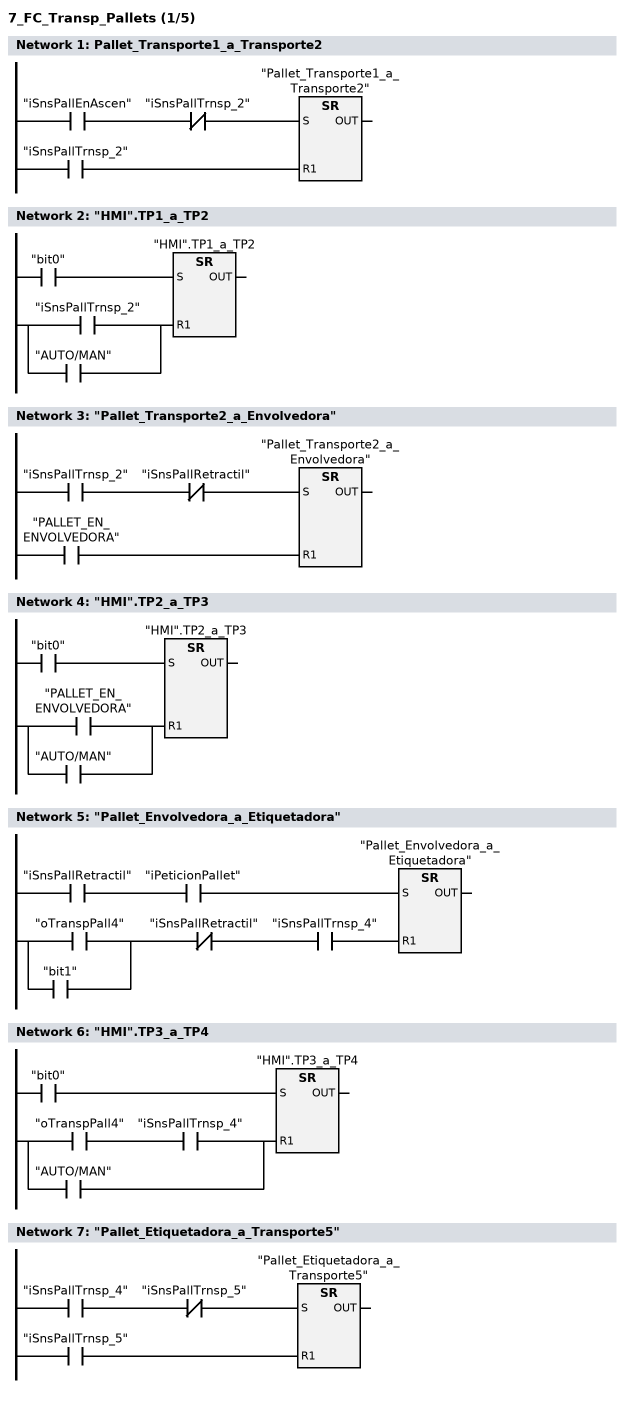
   RUNG wire#powerrail
      Contact( "iSnsPallEnAscen" )
      I_Contact( "iSnsPallTrnsp_2" )
      S_SR(operand := "Pallet_Transporte1_a_Transporte2", r1 := wire#w1)
   END_RUNG
   RUNG wire#powerrail
      Contact( "iSnsPallTrnsp_2" )
   END_RUNG wire#w1
   // the same network as SCL:
   IF "iSnsPallEnAscen" AND NOT "iSnsPallTrnsp_2" THEN
       "Pallet_Transporte1_a_Transporte2" := TRUE;   // SR flip-flop
   END_IF;
   IF "iSnsPallTrnsp_2" THEN "Pallet_Transporte1_a_Transporte2" := FALSE; END_IF;
END_REGION

REGION Network 2: "HMI".TP1_a_TP2
   RUNG wire#powerrail
      Contact( "bit0" )
      S_SR(operand := "HMI".TP1_a_TP2, r1 := wire#w1)
   END_RUNG
   RUNG wire#powerrail
      Contact( "iSnsPallTrnsp_2" )
   END_RUNG wire#w1
   RUNG wire#powerrail
      Contact( "AUTO/MAN" )
   END_RUNG wire#w1
   // the same network as SCL:
   IF "bit0" THEN
       "HMI".TP1_a_TP2 := TRUE;   // SR flip-flop
   END_IF;
   IF "iSnsPallTrnsp_2" OR "AUTO/MAN" THEN "HMI".TP1_a_TP2 := FALSE; END_IF;
END_REGION

REGION Network 3: "Pallet_Transporte2_a_Envolvedora"
   RUNG wire#powerrail
      Contact( "iSnsPallTrnsp_2" )
      I_Contact( "iSnsPallRetractil" )
      S_SR(operand := "Pallet_Transporte2_a_Envolvedora", r1 := wire#w1)
   END_RUNG
   RUNG wire#powerrail
      Contact( "PALLET_EN_ENVOLVEDORA" )
   END_RUNG wire#w1
   // the same network as SCL:
   IF "iSnsPallTrnsp_2" AND NOT "iSnsPallRetractil" THEN
       "Pallet_Transporte2_a_Envolvedora" := TRUE;   // SR flip-flop
   END_IF;
   IF "PALLET_EN_ENVOLVEDORA" THEN "Pallet_Transporte2_a_Envolvedora" := FALSE; END_IF;
END_REGION

REGION Network 4: "HMI".TP2_a_TP3
   RUNG wire#powerrail
      Contact( "bit0" )
      S_SR(operand := "HMI".TP2_a_TP3, r1 := wire#w1)
   END_RUNG
   RUNG wire#powerrail
      Contact( "PALLET_EN_ENVOLVEDORA" )
   END_RUNG wire#w1
   RUNG wire#powerrail
      Contact( "AUTO/MAN" )
   END_RUNG wire#w1
   // the same network as SCL:
   IF "bit0" THEN
       "HMI".TP2_a_TP3 := TRUE;   // SR flip-flop
   END_IF;
   IF "PALLET_EN_ENVOLVEDORA" OR "AUTO/MAN" THEN "HMI".TP2_a_TP3 := FALSE; END_IF;
END_REGION

REGION Network 5: "Pallet_Envolvedora_a_Etiquetadora"
   RUNG wire#powerrail
      Contact( "iSnsPallRetractil" )
      Contact( "iPeticionPallet" )
      S_SR(operand := "Pallet_Envolvedora_a_Etiquetadora", r1 := wire#w2)
   END_RUNG
   RUNG wire#powerrail
      Contact( "oTranspPall4" )
      wire#w1
      I_Contact( "iSnsPallRetractil" )
      Contact( "iSnsPallTrnsp_4" )
   END_RUNG wire#w2
   RUNG wire#powerrail
      Contact( "bit1" )
   END_RUNG wire#w1
   // the same network as SCL:
   IF "iSnsPallRetractil" AND "iPeticionPallet" THEN
       "Pallet_Envolvedora_a_Etiquetadora" := TRUE;   // SR flip-flop
   END_IF;
   IF ("oTranspPall4" OR "bit1") AND NOT "iSnsPallRetractil" AND "iSnsPallTrnsp_4" THEN
       "Pallet_Envolvedora_a_Etiquetadora" := FALSE;
   END_IF;
END_REGION

REGION Network 6: "HMI".TP3_a_TP4
   RUNG wire#powerrail
      Contact( "bit0" )
      S_SR(operand := "HMI".TP3_a_TP4, r1 := wire#w1)
   END_RUNG
   RUNG wire#powerrail
      Contact( "oTranspPall4" )
      Contact( "iSnsPallTrnsp_4" )
   END_RUNG wire#w1
   RUNG wire#powerrail
      Contact( "AUTO/MAN" )
   END_RUNG wire#w1
   // the same network as SCL:
   IF "bit0" THEN
       "HMI".TP3_a_TP4 := TRUE;   // SR flip-flop
   END_IF;
   IF ("oTranspPall4" AND "iSnsPallTrnsp_4") OR "AUTO/MAN" THEN "HMI".TP3_a_TP4 := FALSE; END_IF;
END_REGION

REGION Network 7: "Pallet_Etiquetadora_a_Transporte5"
   RUNG wire#powerrail
      Contact( "iSnsPallTrnsp_4" )
      I_Contact( "iSnsPallTrnsp_5" )
      S_SR(operand := "Pallet_Etiquetadora_a_Transporte5", r1 := wire#w1)
   END_RUNG
   RUNG wire#powerrail
      Contact( "iSnsPallTrnsp_5" )
   END_RUNG wire#w1
   // the same network as SCL:
   IF "iSnsPallTrnsp_4" AND NOT "iSnsPallTrnsp_5" THEN
       "Pallet_Etiquetadora_a_Transporte5" := TRUE;   // SR flip-flop
   END_IF;
   IF "iSnsPallTrnsp_5" THEN "Pallet_Etiquetadora_a_Transporte5" := FALSE; END_IF;
END_REGION

REGION Network 8: "HMI".TP4_a_TP5
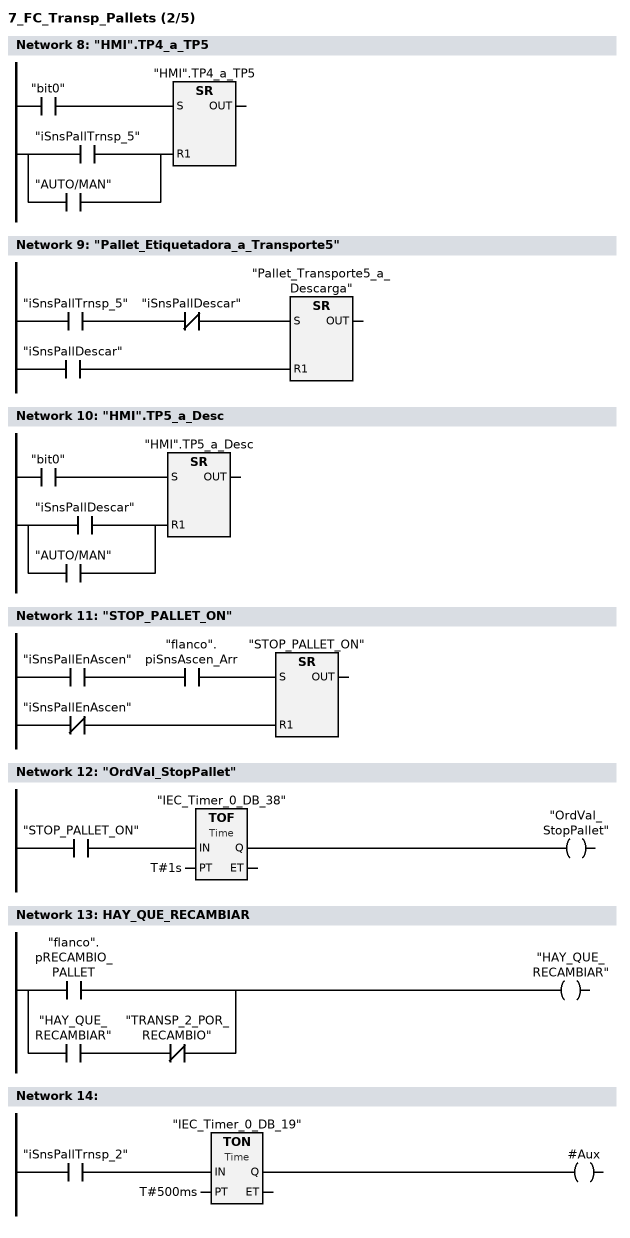
   RUNG wire#powerrail
      Contact( "bit0" )
      S_SR(operand := "HMI".TP4_a_TP5, r1 := wire#w1)
   END_RUNG
   RUNG wire#powerrail
      Contact( "iSnsPallTrnsp_5" )
   END_RUNG wire#w1
   RUNG wire#powerrail
      Contact( "AUTO/MAN" )
   END_RUNG wire#w1
   // the same network as SCL:
   IF "bit0" THEN
       "HMI".TP4_a_TP5 := TRUE;   // SR flip-flop
   END_IF;
   IF "iSnsPallTrnsp_5" OR "AUTO/MAN" THEN "HMI".TP4_a_TP5 := FALSE; END_IF;
END_REGION

REGION Network 9: "Pallet_Etiquetadora_a_Transporte5"
   RUNG wire#powerrail
      Contact( "iSnsPallTrnsp_5" )
      I_Contact( "iSnsPallDescar" )
      S_SR(operand := "Pallet_Transporte5_a_Descarga", r1 := wire#w1)
   END_RUNG
   RUNG wire#powerrail
      Contact( "iSnsPallDescar" )
   END_RUNG wire#w1
   // the same network as SCL:
   IF "iSnsPallTrnsp_5" AND NOT "iSnsPallDescar" THEN
       "Pallet_Transporte5_a_Descarga" := TRUE;   // SR flip-flop
   END_IF;
   IF "iSnsPallDescar" THEN "Pallet_Transporte5_a_Descarga" := FALSE; END_IF;
END_REGION

REGION Network 10: "HMI".TP5_a_Desc
   RUNG wire#powerrail
      Contact( "bit0" )
      S_SR(operand := "HMI".TP5_a_Desc, r1 := wire#w1)
   END_RUNG
   RUNG wire#powerrail
      Contact( "iSnsPallDescar" )
   END_RUNG wire#w1
   RUNG wire#powerrail
      Contact( "AUTO/MAN" )
   END_RUNG wire#w1
   // the same network as SCL:
   IF "bit0" THEN
       "HMI".TP5_a_Desc := TRUE;   // SR flip-flop
   END_IF;
   IF "iSnsPallDescar" OR "AUTO/MAN" THEN "HMI".TP5_a_Desc := FALSE; END_IF;
END_REGION

REGION Network 11: "STOP_PALLET_ON"
   RUNG wire#powerrail
      Contact( "iSnsPallEnAscen" )
      Contact( "flanco".piSnsAscen_Arr )
      S_SR(operand := "STOP_PALLET_ON", r1 := wire#w1)
   END_RUNG
   RUNG wire#powerrail
      I_Contact( "iSnsPallEnAscen" )
   END_RUNG wire#w1
   // the same network as SCL:
   IF "iSnsPallEnAscen" AND "flanco".piSnsAscen_Arr THEN
       "STOP_PALLET_ON" := TRUE;   // SR flip-flop
   END_IF;
   IF NOT "iSnsPallEnAscen" THEN "STOP_PALLET_ON" := FALSE; END_IF;
END_REGION

REGION Network 12: "OrdVal_StopPallet"
   "IEC_Timer_0_DB_38".TOF(in := "STOP_PALLET_ON", pt := T#1s);
   "OrdVal_StopPallet" := "IEC_Timer_0_DB_38".q;
END_REGION

REGION Network 13: HAY_QUE_RECAMBIAR
   RUNG wire#powerrail
      Contact( "flanco".pRECAMBIO_PALLET )
      wire#w1
      Coil( "HAY_QUE_RECAMBIAR" )
   END_RUNG
   RUNG wire#powerrail
      Contact( "HAY_QUE_RECAMBIAR" )
      I_Contact( "TRANSP_2_POR_RECAMBIO" )
   END_RUNG wire#w1
   // the same network as SCL:
   "HAY_QUE_RECAMBIAR" := "flanco".pRECAMBIO_PALLET OR ("HAY_QUE_RECAMBIAR" AND NOT "TRANSP_2_POR_RECAMBIO");
END_REGION

REGION Network 14
   "IEC_Timer_0_DB_19".TON(in := "iSnsPallTrnsp_2", pt := T#500ms);
   #Aux := "IEC_Timer_0_DB_19".q;
END_REGION

REGION Network 15: "TRANSP_2_POR_RECAMBIO"
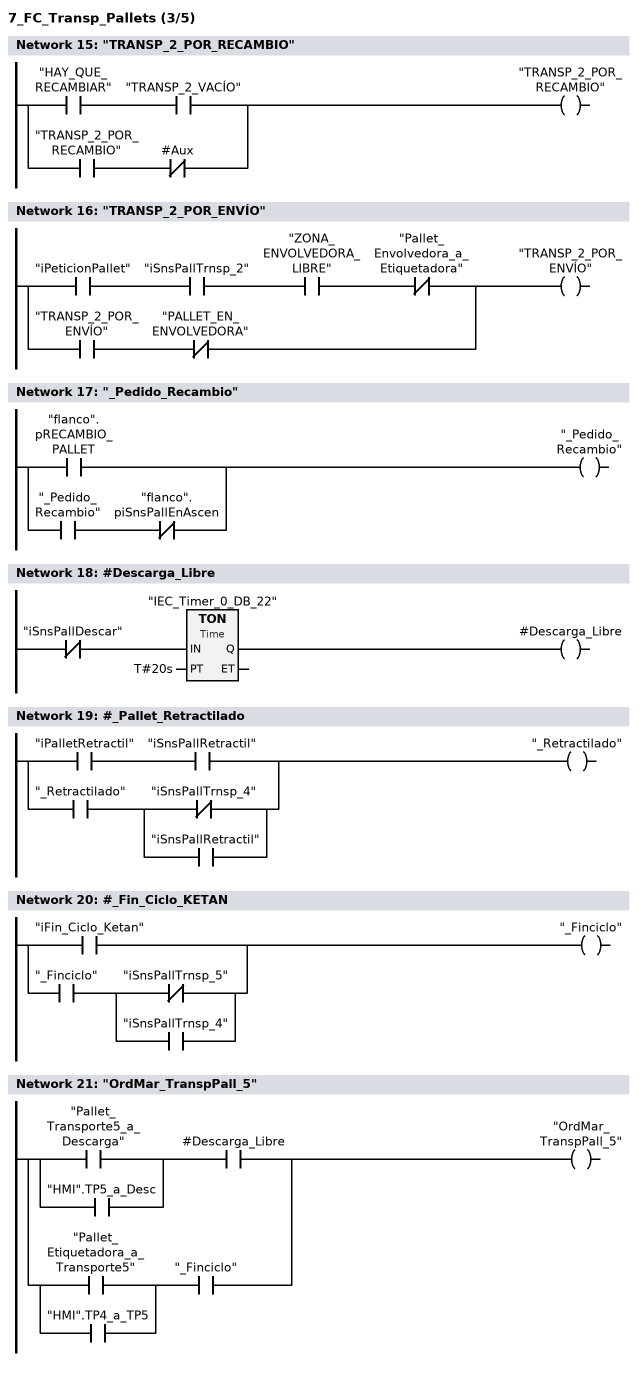
   RUNG wire#powerrail
      Contact( "HAY_QUE_RECAMBIAR" )
      Contact( "TRANSP_2_VACÍO" )
      wire#w1
      Coil( "TRANSP_2_POR_RECAMBIO" )
   END_RUNG
   RUNG wire#powerrail
      Contact( "TRANSP_2_POR_RECAMBIO" )
      I_Contact( #Aux )
   END_RUNG wire#w1
   // the same network as SCL:
   "TRANSP_2_POR_RECAMBIO" := ("HAY_QUE_RECAMBIAR" AND "TRANSP_2_VACÍO") OR ("TRANSP_2_POR_RECAMBIO" AND NOT #Aux);
END_REGION

REGION Network 16: "TRANSP_2_POR_ENVÍO"
   RUNG wire#powerrail
      Contact( "iPeticionPallet" )
      Contact( "iSnsPallTrnsp_2" )
      Contact( "ZONA_ENVOLVEDORA_LIBRE" )
      I_Contact( "Pallet_Envolvedora_a_Etiquetadora" )
      wire#w1
      Coil( "TRANSP_2_POR_ENVÍO" )
   END_RUNG
   RUNG wire#powerrail
      Contact( "TRANSP_2_POR_ENVÍO" )
      I_Contact( "PALLET_EN_ENVOLVEDORA" )
   END_RUNG wire#w1
   // the same network as SCL:
   "TRANSP_2_POR_ENVÍO" := ("iPeticionPallet" AND "iSnsPallTrnsp_2" AND "ZONA_ENVOLVEDORA_LIBRE" AND NOT "Pallet_Envolvedora_a_Etiquetadora") OR ("TRANSP_2_POR_ENVÍO" AND NOT "PALLET_EN_ENVOLVEDORA");
END_REGION

REGION Network 17: "_Pedido_Recambio"
   RUNG wire#powerrail
      Contact( "flanco".pRECAMBIO_PALLET )
      wire#w1
      Coil( "_Pedido_Recambio" )
   END_RUNG
   RUNG wire#powerrail
      Contact( "_Pedido_Recambio" )
      I_Contact( "flanco".piSnsPallEnAscen )
   END_RUNG wire#w1
   // the same network as SCL:
   "_Pedido_Recambio" := "flanco".pRECAMBIO_PALLET OR ("_Pedido_Recambio" AND NOT "flanco".piSnsPallEnAscen);
END_REGION

REGION Network 18: #Descarga_Libre
   "IEC_Timer_0_DB_22".TON(in := NOT "iSnsPallDescar", pt := T#20s);
   #Descarga_Libre := "IEC_Timer_0_DB_22".q;
END_REGION

REGION Network 19: #_Pallet_Retractilado
   RUNG wire#powerrail
      Contact( "iPalletRetractil" )
      Contact( "iSnsPallRetractil" )
      wire#w1
      Coil( "_Retractilado" )
   END_RUNG
   RUNG wire#powerrail
      Contact( "_Retractilado" )
      wire#w2
      I_Contact( "iSnsPallTrnsp_4" )
   END_RUNG wire#w1
   RUNG wire#w2
      Contact( "iSnsPallRetractil" )
   END_RUNG wire#w1
   // the same network as SCL:
   "_Retractilado" := ("iPalletRetractil" AND "iSnsPallRetractil") OR ("_Retractilado" AND (NOT "iSnsPallTrnsp_4" OR "iSnsPallRetractil"));
END_REGION

REGION Network 20: #_Fin_Ciclo_KETAN
   RUNG wire#powerrail
      Contact( "iFin_Ciclo_Ketan" )
      wire#w1
      Coil( "_Finciclo" )
   END_RUNG
   RUNG wire#powerrail
      Contact( "_Finciclo" )
      wire#w2
      I_Contact( "iSnsPallTrnsp_5" )
   END_RUNG wire#w1
   RUNG wire#w2
      Contact( "iSnsPallTrnsp_4" )
   END_RUNG wire#w1
   // the same network as SCL:
   "_Finciclo" := "iFin_Ciclo_Ketan" OR ("_Finciclo" AND (NOT "iSnsPallTrnsp_5" OR "iSnsPallTrnsp_4"));
END_REGION

REGION Network 21: "OrdMar_TranspPall_5"
   RUNG wire#powerrail
      Contact( "Pallet_Transporte5_a_Descarga" )
      wire#w1
      Contact( #Descarga_Libre )
      wire#w2
      Coil( "OrdMar_TranspPall_5" )
   END_RUNG
   RUNG wire#powerrail
      Contact( "HMI".TP5_a_Desc )
   END_RUNG wire#w1
   RUNG wire#powerrail
      Contact( "Pallet_Etiquetadora_a_Transporte5" )
      wire#w3
      Contact( "_Finciclo" )
   END_RUNG wire#w2
   RUNG wire#powerrail
      Contact( "HMI".TP4_a_TP5 )
   END_RUNG wire#w3
   // the same network as SCL:
   "OrdMar_TranspPall_5" := (("Pallet_Transporte5_a_Descarga" OR "HMI".TP5_a_Desc) AND #Descarga_Libre) OR (("Pallet_Etiquetadora_a_Transporte5" OR "HMI".TP4_a_TP5) AND "_Finciclo");
END_REGION

REGION Network 22: "OrdMar_TranspPall_4"
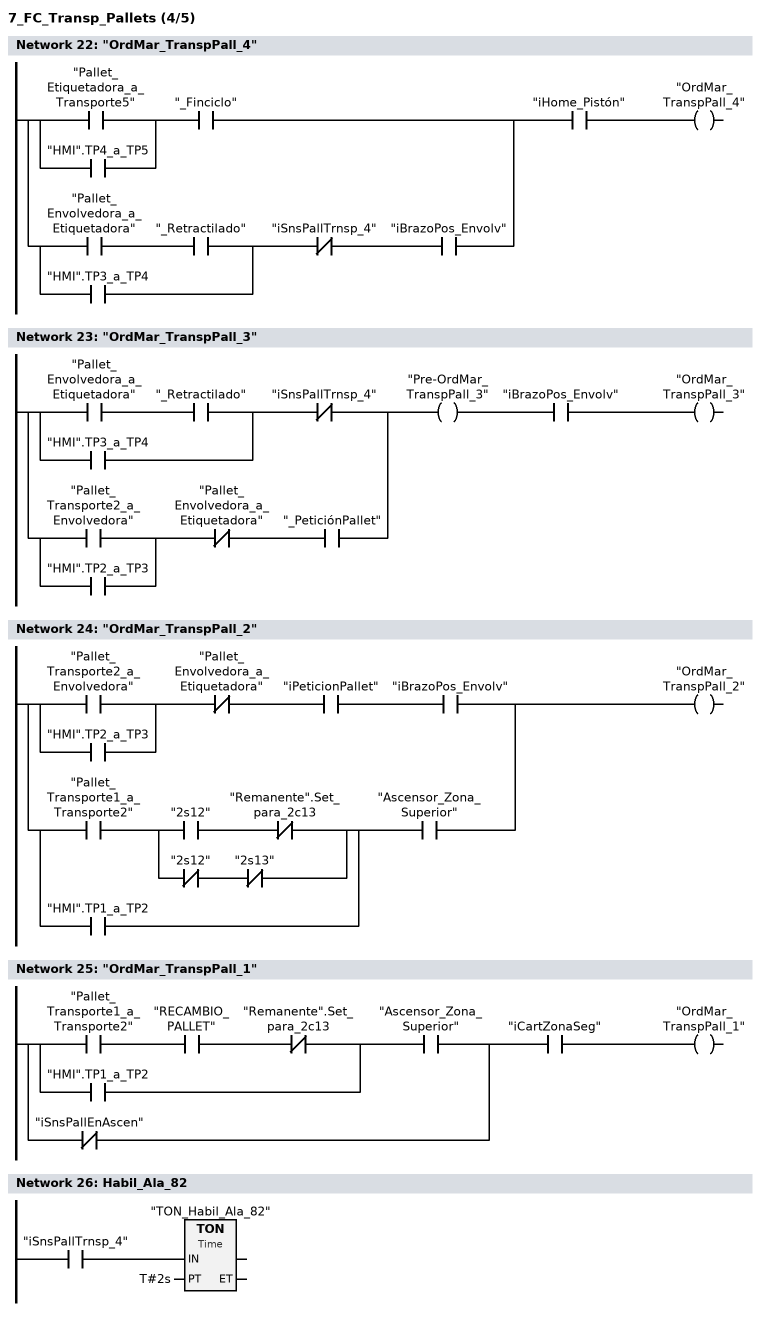
   RUNG wire#powerrail
      Contact( "Pallet_Etiquetadora_a_Transporte5" )
      wire#w1
      Contact( "_Finciclo" )
      wire#w2
      Contact( "iHome_Pistón" )
      Coil( "OrdMar_TranspPall_4" )
   END_RUNG
   RUNG wire#powerrail
      Contact( "HMI".TP4_a_TP5 )
   END_RUNG wire#w1
   RUNG wire#powerrail
      Contact( "Pallet_Envolvedora_a_Etiquetadora" )
      Contact( "_Retractilado" )
      wire#w3
      I_Contact( "iSnsPallTrnsp_4" )
      Contact( "iBrazoPos_Envolv" )
   END_RUNG wire#w2
   RUNG wire#powerrail
      Contact( "HMI".TP3_a_TP4 )
   END_RUNG wire#w3
   // the same network as SCL:
   "OrdMar_TranspPall_4" := ((("Pallet_Etiquetadora_a_Transporte5" OR "HMI".TP4_a_TP5) AND "_Finciclo") OR ((("Pallet_Envolvedora_a_Etiquetadora" AND "_Retractilado") OR "HMI".TP3_a_TP4) AND NOT "iSnsPallTrnsp_4" AND "iBrazoPos_Envolv")) AND "iHome_Pistón";
END_REGION

REGION Network 23: "OrdMar_TranspPall_3"
   RUNG wire#powerrail
      Contact( "Pallet_Envolvedora_a_Etiquetadora" )
      Contact( "_Retractilado" )
      wire#w1
      I_Contact( "iSnsPallTrnsp_4" )
      wire#w2
      Coil( "Pre-OrdMar_TranspPall_3" )
      Contact( "iBrazoPos_Envolv" )
      Coil( "OrdMar_TranspPall_3" )
   END_RUNG
   RUNG wire#powerrail
      Contact( "HMI".TP3_a_TP4 )
   END_RUNG wire#w1
   RUNG wire#powerrail
      Contact( "Pallet_Transporte2_a_Envolvedora" )
      wire#w3
      I_Contact( "Pallet_Envolvedora_a_Etiquetadora" )
      Contact( "_PeticiónPallet" )
   END_RUNG wire#w2
   RUNG wire#powerrail
      Contact( "HMI".TP2_a_TP3 )
   END_RUNG wire#w3
   // the same network as SCL:
   "Pre-OrdMar_TranspPall_3" := ((("Pallet_Envolvedora_a_Etiquetadora" AND "_Retractilado") OR "HMI".TP3_a_TP4) AND NOT "iSnsPallTrnsp_4") OR (("Pallet_Transporte2_a_Envolvedora" OR "HMI".TP2_a_TP3) AND NOT "Pallet_Envolvedora_a_Etiquetadora" AND "_PeticiónPallet");
   "OrdMar_TranspPall_3" := "Pre-OrdMar_TranspPall_3" AND "iBrazoPos_Envolv";
END_REGION

REGION Network 24: "OrdMar_TranspPall_2"
   RUNG wire#powerrail
      Contact( "Pallet_Transporte2_a_Envolvedora" )
      wire#w1
      I_Contact( "Pallet_Envolvedora_a_Etiquetadora" )
      Contact( "iPeticionPallet" )
      Contact( "iBrazoPos_Envolv" )
      wire#w2
      Coil( "OrdMar_TranspPall_2" )
   END_RUNG
   RUNG wire#powerrail
      Contact( "HMI".TP2_a_TP3 )
   END_RUNG wire#w1
   RUNG wire#powerrail
      Contact( "Pallet_Transporte1_a_Transporte2" )
      wire#w3
      Contact( "2s12" )
      I_Contact( "Remanente".Set_para_2c13 )
      wire#w4
      Contact( "Ascensor_Zona_Superior" )
   END_RUNG wire#w2
   RUNG wire#w3
      I_Contact( "2s12" )
      I_Contact( "2s13" )
   END_RUNG wire#w4
   RUNG wire#powerrail
      Contact( "HMI".TP1_a_TP2 )
   END_RUNG wire#w4
   // the same network as SCL:
   "OrdMar_TranspPall_2" := (("Pallet_Transporte2_a_Envolvedora" OR "HMI".TP2_a_TP3) AND NOT "Pallet_Envolvedora_a_Etiquetadora" AND "iPeticionPallet" AND "iBrazoPos_Envolv") OR ((("Pallet_Transporte1_a_Transporte2" AND (("2s12" AND NOT "Remanente".Set_para_2c13) OR (NOT "2s12" AND NOT "2s13"))) OR "HMI".TP1_a_TP2) AND "Ascensor_Zona_Superior");
END_REGION

REGION Network 25: "OrdMar_TranspPall_1"
   RUNG wire#powerrail
      Contact( "Pallet_Transporte1_a_Transporte2" )
      Contact( "RECAMBIO_PALLET" )
      I_Contact( "Remanente".Set_para_2c13 )
      wire#w1
      Contact( "Ascensor_Zona_Superior" )
      wire#w2
      Contact( "iCartZonaSeg" )
      Coil( "OrdMar_TranspPall_1" )
   END_RUNG
   RUNG wire#powerrail
      Contact( "HMI".TP1_a_TP2 )
   END_RUNG wire#w1
   RUNG wire#powerrail
      I_Contact( "iSnsPallEnAscen" )
   END_RUNG wire#w2
   // the same network as SCL:
   "OrdMar_TranspPall_1" := (((("Pallet_Transporte1_a_Transporte2" AND "RECAMBIO_PALLET" AND NOT "Remanente".Set_para_2c13) OR "HMI".TP1_a_TP2) AND "Ascensor_Zona_Superior") OR NOT "iSnsPallEnAscen") AND "iCartZonaSeg";
END_REGION

REGION Network 26: Habil_Ala_82
   "TON_Habil_Ala_82".TON(IN := "iSnsPallTrnsp_4", PT := T#2s);
END_REGION

REGION Network 27: Habil_Ala_82 (Cont.)
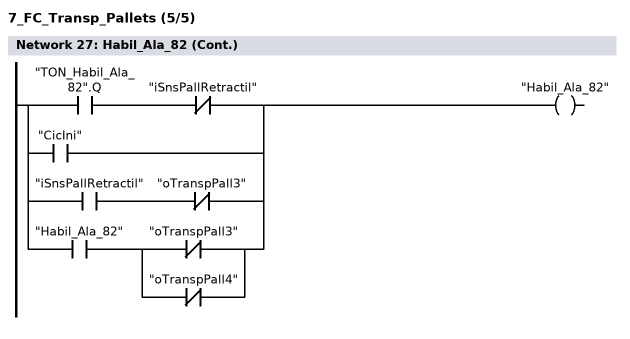
   RUNG wire#powerrail
      Contact( "TON_Habil_Ala_82".Q )
      I_Contact( "iSnsPallRetractil" )
      wire#w1
      Coil( "Habil_Ala_82" )
   END_RUNG
   RUNG wire#powerrail
      Contact( "CicIni" )
   END_RUNG wire#w1
   RUNG wire#powerrail
      Contact( "iSnsPallRetractil" )
      I_Contact( "oTranspPall3" )
   END_RUNG wire#w1
   RUNG wire#powerrail
      Contact( "Habil_Ala_82" )
      wire#w2
      I_Contact( "oTranspPall3" )
   END_RUNG wire#w1
   RUNG wire#w2
      I_Contact( "oTranspPall4" )
   END_RUNG wire#w1
   // the same network as SCL:
   "Habil_Ala_82" := ("TON_Habil_Ala_82".Q AND NOT "iSnsPallRetractil") OR "CicIni" OR ("iSnsPallRetractil" AND NOT "oTranspPall3") OR ("Habil_Ala_82" AND (NOT "oTranspPall3" OR NOT "oTranspPall4"));
END_REGION
END_FUNCTION

FUNCTION "8_FC_Almacen_Pallets" : Void   // FC15, LAD
{ S7_Optimized_Access := 'FALSE' }
VERSION : 0.1
BEGIN

REGION Network 1: #Aux
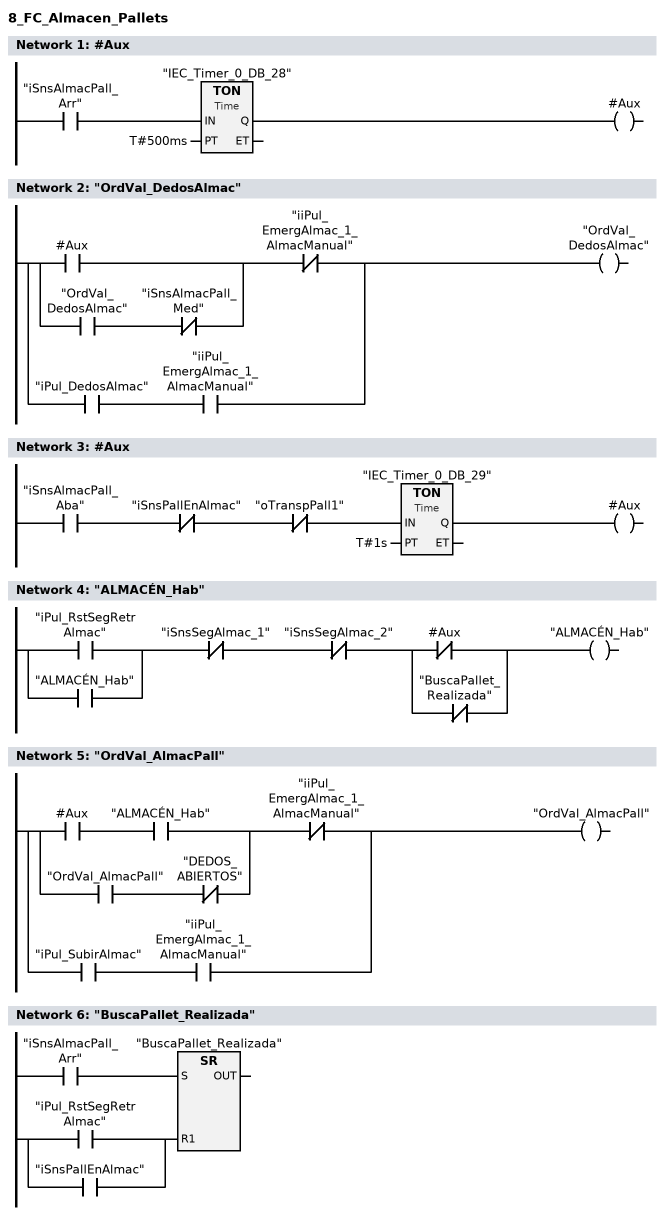
   "IEC_Timer_0_DB_28".TON(in := "iSnsAlmacPall_Arr", pt := T#500ms);
   #Aux := "IEC_Timer_0_DB_28".q;
END_REGION

REGION Network 2: "OrdVal_DedosAlmac"
   RUNG wire#powerrail
      Contact( #Aux )
      wire#w1
      I_Contact( "iiPul_EmergAlmac_1_AlmacManual" )
      wire#w2
      Coil( "OrdVal_DedosAlmac" )
   END_RUNG
   RUNG wire#powerrail
      Contact( "OrdVal_DedosAlmac" )
      I_Contact( "iSnsAlmacPall_Med" )
   END_RUNG wire#w1
   RUNG wire#powerrail
      Contact( "iPul_DedosAlmac" )
      Contact( "iiPul_EmergAlmac_1_AlmacManual" )
   END_RUNG wire#w2
   // the same network as SCL:
   "OrdVal_DedosAlmac" := ((#Aux OR ("OrdVal_DedosAlmac" AND NOT "iSnsAlmacPall_Med")) AND NOT "iiPul_EmergAlmac_1_AlmacManual") OR ("iPul_DedosAlmac" AND "iiPul_EmergAlmac_1_AlmacManual");
END_REGION

REGION Network 3: #Aux
   "IEC_Timer_0_DB_29".TON(IN := "iSnsAlmacPall_Aba" AND NOT "iSnsPallEnAlmac" AND NOT "oTranspPall1",
                           PT := T#1s);
   #Aux := "IEC_Timer_0_DB_29".Q;
END_REGION

REGION Network 4: "ALMACÉN_Hab"
   RUNG wire#powerrail
      Contact( "iPul_RstSegRetrAlmac" )
      wire#w1
      I_Contact( "iSnsSegAlmac_1" )
      I_Contact( "iSnsSegAlmac_2" )
      wire#w2
      I_Contact( #Aux )
      wire#w3
      Coil( "ALMACÉN_Hab" )
   END_RUNG
   RUNG wire#powerrail
      Contact( "ALMACÉN_Hab" )
   END_RUNG wire#w1
   RUNG wire#w2
      I_Contact( "BuscaPallet_Realizada" )
   END_RUNG wire#w3
   // the same network as SCL:
   "ALMACÉN_Hab" := ("iPul_RstSegRetrAlmac" OR "ALMACÉN_Hab") AND NOT "iSnsSegAlmac_1" AND NOT "iSnsSegAlmac_2" AND (NOT #Aux OR NOT "BuscaPallet_Realizada");
END_REGION

REGION Network 5: "OrdVal_AlmacPall"
   RUNG wire#powerrail
      Contact( #Aux )
      Contact( "ALMACÉN_Hab" )
      wire#w1
      I_Contact( "iiPul_EmergAlmac_1_AlmacManual" )
      wire#w2
      Coil( "OrdVal_AlmacPall" )
   END_RUNG
   RUNG wire#powerrail
      Contact( "OrdVal_AlmacPall" )
      I_Contact( "DEDOS_ABIERTOS" )
   END_RUNG wire#w1
   RUNG wire#powerrail
      Contact( "iPul_SubirAlmac" )
      Contact( "iiPul_EmergAlmac_1_AlmacManual" )
   END_RUNG wire#w2
   // the same network as SCL:
   "OrdVal_AlmacPall" := (((#Aux AND "ALMACÉN_Hab") OR ("OrdVal_AlmacPall" AND NOT "DEDOS_ABIERTOS")) AND NOT "iiPul_EmergAlmac_1_AlmacManual") OR ("iPul_SubirAlmac" AND "iiPul_EmergAlmac_1_AlmacManual");
END_REGION

REGION Network 6: "BuscaPallet_Realizada"
   RUNG wire#powerrail
      Contact( "iSnsAlmacPall_Arr" )
      S_SR(operand := "BuscaPallet_Realizada", r1 := wire#w1)
   END_RUNG
   RUNG wire#powerrail
      Contact( "iPul_RstSegRetrAlmac" )
   END_RUNG wire#w1
   RUNG wire#powerrail
      Contact( "iSnsPallEnAlmac" )
   END_RUNG wire#w1
   // the same network as SCL:
   IF "iSnsAlmacPall_Arr" THEN
       "BuscaPallet_Realizada" := TRUE;   // SR flip-flop
   END_IF;
   IF "iPul_RstSegRetrAlmac" OR "iSnsPallEnAlmac" THEN "BuscaPallet_Realizada" := FALSE; END_IF;
END_REGION
END_FUNCTION

FUNCTION "10_ELEMENTO_HH" : Void   // FC28, LAD
{ S7_Optimized_Access := 'FALSE' }
VERSION : 0.1
// En viada la primer caja, se encarga de acomodarla y enviar la segunda
BEGIN

REGION Network 1: ESTADO ACTIVO
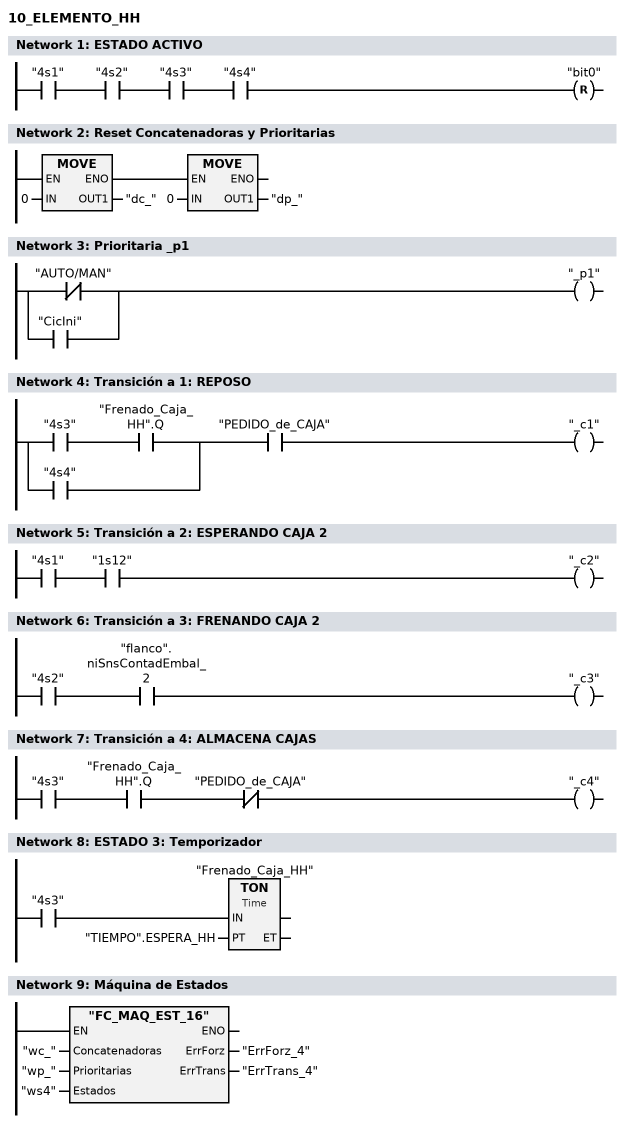
   RUNG wire#powerrail
      Contact( "4s1" )
      Contact( "4s2" )
      Contact( "4s3" )
      Contact( "4s4" )
      R_Coil( "bit0" )
   END_RUNG
   // the same network as SCL:
   IF "4s1" AND "4s2" AND "4s3" AND "4s4" THEN "bit0" := FALSE; END_IF;
END_REGION

REGION Network 2: Reset Concatenadoras y Prioritarias
   RUNG wire#powerrail
      { S7_GenerateENO := "TRUE" } Move(in := 0, out1 => "dc_")
      { S7_GenerateENO := "TRUE" } Move(in := 0, out1 => "dp_")
   END_RUNG
   // the same network as SCL:
   // ENO of a box is taken as its EN; it also drops when the box reports an error
   "dc_" := 0;
   "dp_" := 0;
END_REGION

REGION Network 3: Prioritaria _p1
   RUNG wire#powerrail
      I_Contact( "AUTO/MAN" )
      wire#w1
      Coil( "_p1" )
   END_RUNG
   RUNG wire#powerrail
      Contact( "CicIni" )
   END_RUNG wire#w1
   // the same network as SCL:
   "_p1" := NOT "AUTO/MAN" OR "CicIni";
END_REGION

REGION Network 4: Transición a 1: REPOSO
   RUNG wire#powerrail
      Contact( "4s3" )
      Contact( "Frenado_Caja_HH".Q )
      wire#w1
      Contact( "PEDIDO_de_CAJA" )
      Coil( "_c1" )
   END_RUNG
   RUNG wire#powerrail
      Contact( "4s4" )
   END_RUNG wire#w1
   // the same network as SCL:
   "_c1" := (("4s3" AND "Frenado_Caja_HH".Q) OR "4s4") AND "PEDIDO_de_CAJA";
END_REGION

REGION Network 5: Transición a 2: ESPERANDO CAJA 2
   RUNG wire#powerrail
      Contact( "4s1" )
      Contact( "1s12" )
      Coil( "_c2" )
   END_RUNG
   // the same network as SCL:
   "_c2" := "4s1" AND "1s12";
END_REGION

REGION Network 6: Transición a 3: FRENANDO CAJA 2
   RUNG wire#powerrail
      Contact( "4s2" )
      Contact( "flanco".niSnsContadEmbal_2 )
      Coil( "_c3" )
   END_RUNG
   // the same network as SCL:
   "_c3" := "4s2" AND "flanco".niSnsContadEmbal_2;
END_REGION

REGION Network 7: Transición a 4: ALMACENA CAJAS
   RUNG wire#powerrail
      Contact( "4s3" )
      Contact( "Frenado_Caja_HH".Q )
      I_Contact( "PEDIDO_de_CAJA" )
      Coil( "_c4" )
   END_RUNG
   // the same network as SCL:
   "_c4" := "4s3" AND "Frenado_Caja_HH".Q AND NOT "PEDIDO_de_CAJA";
END_REGION

REGION Network 8: ESTADO 3: Temporizador
   "Frenado_Caja_HH".TON(in := "4s3", pt := "TIEMPO".ESPERA_HH);
END_REGION

REGION Network 9: Máquina de Estados
   RUNG wire#powerrail
      "FC_MAQ_EST_16"(Concatenadoras := "wc_", Prioritarias := "wp_", Estados := "ws4", ErrForz => "ErrForz_4", ErrTrans => "ErrTrans_4")
   END_RUNG
   // the same network as SCL:
   "FC_MAQ_EST_16"(Concatenadoras := "wc_",
                   Prioritarias := "wp_",
                   Estados := "ws4",
                   ErrForz => "ErrForz_4",
                   ErrTrans => "ErrTrans_4");
END_REGION
END_FUNCTION

FUNCTION "11_FC_Cartoneo_Manual" : Void   // FC31, LAD
{ S7_Optimized_Access := 'FALSE' }
VERSION : 0.1
   VAR_TEMP   // added for the SCL form of the ladder/FBD networks
      _w1 : Bool;
      _w2 : Bool;
   END_VAR
BEGIN

REGION Network 1: Habilitación Cartoneo Manual - Desde HMI
END_REGION

REGION Network 2: Freno del ciclo de paletizador
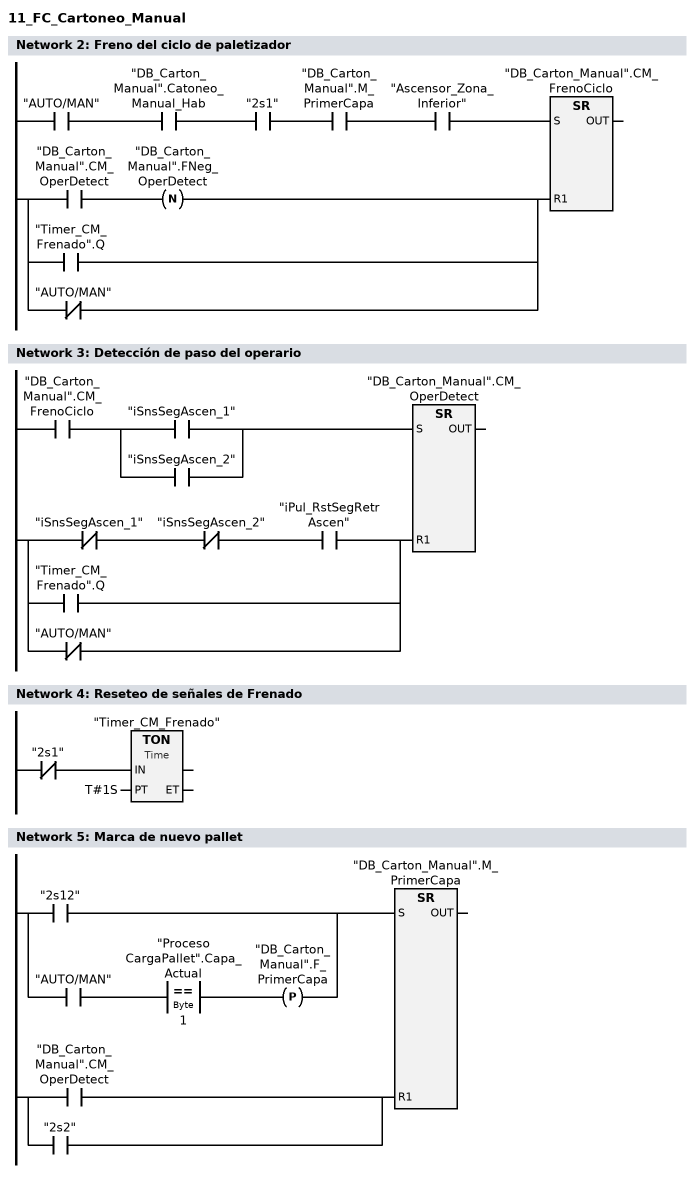
   RUNG wire#powerrail
      Contact( "AUTO/MAN" )
      Contact( "DB_Carton_Manual".Catoneo_Manual_Hab )
      Contact( "2s1" )
      Contact( "DB_Carton_Manual".M_PrimerCapa )
      Contact( "Ascensor_Zona_Inferior" )
      S_SR(operand := "DB_Carton_Manual".CM_FrenoCiclo, r1 := wire#w1)
   END_RUNG
   RUNG wire#powerrail
      Contact( "DB_Carton_Manual".CM_OperDetect )
      N_Trig( "DB_Carton_Manual".FNeg_OperDetect )
   END_RUNG wire#w1
   RUNG wire#powerrail
      Contact( "Timer_CM_Frenado".Q )
   END_RUNG wire#w1
   RUNG wire#powerrail
      I_Contact( "AUTO/MAN" )
   END_RUNG wire#w1
   // the same network as SCL:
   #_w1 := NOT "DB_Carton_Manual".CM_OperDetect AND "DB_Carton_Manual".FNeg_OperDetect;   // falling edge
   "DB_Carton_Manual".FNeg_OperDetect := "DB_Carton_Manual".CM_OperDetect;
   IF "AUTO/MAN" AND "DB_Carton_Manual".Catoneo_Manual_Hab AND "2s1" AND "DB_Carton_Manual".M_PrimerCapa AND "Ascensor_Zona_Inferior" THEN
       "DB_Carton_Manual".CM_FrenoCiclo := TRUE;   // SR flip-flop
   END_IF;
   IF #_w1 OR "Timer_CM_Frenado".Q OR NOT "AUTO/MAN" THEN "DB_Carton_Manual".CM_FrenoCiclo := FALSE; END_IF;
END_REGION

REGION Network 3: Detección de paso del operario
   RUNG wire#powerrail
      Contact( "DB_Carton_Manual".CM_FrenoCiclo )
      wire#w1
      Contact( "iSnsSegAscen_1" )
      wire#w2
      S_SR(operand := "DB_Carton_Manual".CM_OperDetect, r1 := wire#w3)
   END_RUNG
   RUNG wire#w1
      Contact( "iSnsSegAscen_2" )
   END_RUNG wire#w2
   RUNG wire#powerrail
      I_Contact( "iSnsSegAscen_1" )
      I_Contact( "iSnsSegAscen_2" )
      Contact( "iPul_RstSegRetrAscen" )
   END_RUNG wire#w3
   RUNG wire#powerrail
      Contact( "Timer_CM_Frenado".Q )
   END_RUNG wire#w3
   RUNG wire#powerrail
      I_Contact( "AUTO/MAN" )
   END_RUNG wire#w3
   // the same network as SCL:
   IF "DB_Carton_Manual".CM_FrenoCiclo AND ("iSnsSegAscen_1" OR "iSnsSegAscen_2") THEN
       "DB_Carton_Manual".CM_OperDetect := TRUE;   // SR flip-flop
   END_IF;
   IF (NOT "iSnsSegAscen_1" AND NOT "iSnsSegAscen_2" AND "iPul_RstSegRetrAscen") OR "Timer_CM_Frenado".Q OR NOT "AUTO/MAN" THEN
       "DB_Carton_Manual".CM_OperDetect := FALSE;
   END_IF;
END_REGION

REGION Network 4: Reseteo de señales de Frenado
   "Timer_CM_Frenado".TON(IN := NOT "2s1", PT := T#1S);
END_REGION

REGION Network 5: Marca de nuevo pallet
   RUNG wire#powerrail
      Contact( "2s12" )
      wire#w1
      S_SR(operand := "DB_Carton_Manual".M_PrimerCapa, r1 := wire#w2)
   END_RUNG
   RUNG wire#powerrail
      Contact( "AUTO/MAN" )
      { S7_Templates := "SrcType := Byte" } EQ_Contact(in1 := "Proceso CargaPallet".Capa_Actual, in2 := 1)
      P_Trig( "DB_Carton_Manual".F_PrimerCapa )
   END_RUNG wire#w1
   RUNG wire#powerrail
      Contact( "DB_Carton_Manual".CM_OperDetect )
   END_RUNG wire#w2
   RUNG wire#powerrail
      Contact( "2s2" )
   END_RUNG wire#w2
   // the same network as SCL:
   #_w1 := "AUTO/MAN" AND ("Proceso CargaPallet".Capa_Actual = 1);
   #_w2 := #_w1 AND NOT "DB_Carton_Manual".F_PrimerCapa;   // rising edge
   "DB_Carton_Manual".F_PrimerCapa := #_w1;
   IF "2s12" OR #_w2 THEN
       "DB_Carton_Manual".M_PrimerCapa := TRUE;   // SR flip-flop
   END_IF;
   IF "DB_Carton_Manual".CM_OperDetect OR "2s2" THEN "DB_Carton_Manual".M_PrimerCapa := FALSE; END_IF;
END_REGION
END_FUNCTION

// folder: Movimiento DATOS

FUNCTION "FC_ELEM_PROX" : Void   // FC1, STL
{ S7_Optimized_Access := 'FALSE' }
VERSION : 0.1
BEGIN

REGION Network 1: Constantes
         L     "Proceso Dosificador".Cant_Pallets;
         T     #Nro_Pallet;
         L     "Proceso Dosificador".Capa_Actual;
         T     #Capa_Actual;
         L     38;
         T     #Length_Capas;
         L     54;
         T     #Offset_Capas;
         L     6;
         T     #Length_Filas_DB;
         L     0;
         T     #Offset_Filas_DB;
         L     1;
         T     #Length_Elementos_DB_bit;
         L     0;
         T     #Offset_Elementos_DB_bit;

         L     1;
         T     #Índice_Filas;
         T     #Índice_Elementos;

         L     "Puntero".Max_Nro_Elementos;
         T     #Max_Nro_Elementos;
         L     "Puntero".Max_Nro_Filas;
         T     #Max_Nro_Filas;
         L     "Puntero".Max_Nro_Capas;
         T     #Max_Nro_Capas;
END_REGION

REGION Network 2: Adress_Capa
         L     #Capa_Actual;
         L     1;
         -I;
         L     #Length_Capas;
         *I;
         L     #Offset_Capas;
         +I;
         T     #Adress_Capa;
END_REGION

REGION Network 3: Adress_Filas
   New_Fil:NOP   0;
         L     #Índice_Filas;
         L     1;
         -I;
         L     #Length_Filas_DB;
         *I;
         L     #Offset_Filas_DB;
         +I;
         L     #Adress_Capa;
         +I;
         SLD   3;
         T     #Adress_Filas_DB_bit;
END_REGION

REGION Network 4: Adress_Elementos_DB
   New_Ele:NOP   0;
         L     #Índice_Elementos;
         L     1;
         -I;
         L     #Length_Elementos_DB_bit;
         *I;
         L     #Offset_Elementos_DB_bit;
         +I;
         L     #Adress_Filas_DB_bit;
         +I;
         T     #Adress_Elementos_DB_bit;
END_REGION

REGION Network 5: AR1
         L     #Adress_Elementos_DB_bit;
         LAR1;
END_REGION

REGION Network 6: Habilita ir 1 lugar a la IZQ
         OPN   "DB_Receta_Actual";
         SET;
         R     #Habil_1_IZQ;
         L     #Índice_Elementos;
         L     #Max_Nro_Elementos;
         >=I;
         JC    No1IZQ;
         TAR1  AR2;
         L     1;
         +AR2;
         O     DBX [ AR2 , P#0.0 ];
         O     DBX [ AR2 , P#2.0 ];
         =     #Habil_1_IZQ;
   No1IZQ:NOP   0;
END_REGION

REGION Network 7: Habilita ir 2 lugar a la IZQ
         OPN   "DB_Receta_Actual";
         SET;
         R     #Habil_2_IZQ;
         L     #Índice_Elementos;
         L     1;
         +I;
         L     #Max_Nro_Elementos;
         >=I;
         JC    No2IZQ;
         TAR1  AR2;
         L     2;
         +AR2;
         O     DBX [ AR2 , P#0.0 ];
         O     DBX [ AR2 , P#2.0 ];
         =     #Habil_2_IZQ;
   No2IZQ:NOP   0;
END_REGION

REGION Network 8: Habilita ir a ABA_Elem_1
         OPN   "DB_Receta_Actual";
         SET;
         R     #Habil_1_ABA;
         L     #Índice_Filas;
         L     #Max_Nro_Filas;
         >=I;
         JC    No1ABA;
         L     #Adress_Filas_DB_bit;
         SRD   3;
         L     #Length_Filas_DB;
         +I;
         SLD   3;
         L     #Offset_Elementos_DB_bit;
         +I;
         LAR2;
         O     DBX [AR2, P#0.0];
         O     DBX [ AR2 , P#2.0 ];
         =     #Habil_1_ABA;
   No1ABA:NOP   0;
END_REGION

REGION Network 9: Habilita ir a ABA_Elem_2
         OPN   "DB_Receta_Actual";
         SET;
         R     #Habil_2_ABA;
         L     #Índice_Filas;
         L     #Max_Nro_Filas;
         >=I;
         JC    No2ABA;
         L     #Adress_Filas_DB_bit;
         SRD   3;
         L     #Length_Filas_DB;
         +I;
         SLD   3;
         L     #Offset_Elementos_DB_bit;
         +I;
         L     #Length_Elementos_DB_bit;
         +I;
         LAR2;
         O     DBX [AR2, P#0.0];
         O     DBX [ AR2 , P#2.0 ];
         =     #Habil_2_ABA;
   No2ABA:NOP   0;
END_REGION

REGION Network 10: Habilita cambiar de CAPA_Elem_1
         OPN   "DB_Receta_Actual";
         SET;
         R     #Habil_1_CAPA;
         L     #Capa_Actual;
         L     #Max_Nro_Capas;
         >=I;
         JC    No1CAPA;
         L     #Adress_Capa;
         L     #Length_Capas;
         +I;
         L     #Offset_Filas_DB;
         +I;
         SLD   3;
         L     #Offset_Elementos_DB_bit;
         +I;
         LAR2;
         O     DBX [AR2, P#0.0];
         O     DBX [ AR2 , P#2.0 ];
         =     #Habil_1_CAPA;
   No1CAPA:NOP   0;
END_REGION
